(* Logix 5000 project; controller FV vendor 1 type 14 code 217 rev 31.11; software revision 31.00; part 9 of 63 *)
(* tags used below, declared in another part *)
   FR_CFG1_P : PlantItem;   // CFG1_P
   FR_CFG1_P_RawInput : ALIAS FOR RIO_Rack_2:12:I.Data.0;   // FR_CFG1_P
   FR_CFG2_P : PlantItem;   // CFG2_P
   FR_CFG2_P_RawInput : ALIAS FOR RIO_Rack_2:12:I.Data.1;   // FR_CFG2_P
   FR_DEFOAMER : PlantItem;   // DEFOAMER
   FR_DEFOAMER_RawInput : ALIAS FOR RIO_Rack_2:4:I.Data.6;   // FR_DEFOAMER
   FR_Delphi_I : DINT[60];
   FR_FV26_ROTO : PlantItem;   // FV26_ROTO
   FR_FV26_ROTO_RawInput : ALIAS FOR RIO_Rack_2:12:I.Data.10;   // FR_FV26_ROTO
   FR_FV27_ROTO : PlantItem;   // FV27_ROTO
   FR_FV27_ROTO_RawInput : ALIAS FOR RIO_Rack_2:12:I.Data.11;   // FR_FV27_ROTO
   FR_FV28_ROTO : PlantItem;   // FV28_ROTO
   FR_FV28_ROTO_RawInput : ALIAS FOR RIO_Rack_2:12:I.Data.12;   // FR_FV28_ROTO
   FR_FV29_ROTO : PlantItem;   // FV29_ROTO
   FR_FV29_ROTO_RawInput : ALIAS FOR RIO_Rack_2:12:I.Data.13;   // FR_FV29_ROTO
   FR_FV30_ROTO : PlantItem;   // FV30_ROTO
   FR_FV30_ROTO_RawInput : ALIAS FOR RIO_Rack_2:12:I.Data.14;   // FR_FV30_ROTO
   FR_FV31_ROTO : PlantItem;   // FV31_ROTO
   FR_FV31_ROTO_RawInput : ALIAS FOR RIO_Rack_2:12:I.Data.15;   // FR_FV31_ROTO
   FR_OXY_SW1 : PlantItem;   // OXY_SW1
   FR_OXY_SW1_RawInput : ALIAS FOR RIO_Rack_2:3:I.Data.28;   // FR_OXY_SW1
   FR_OXY_SW2 : PlantItem;   // OXY_SW2
   FR_OXY_SW2_RawInput : ALIAS FOR RIO_Rack_2:3:I.Data.29;   // FR_OXY_SW2
   FR_PANELESTOP : PlantItem;   // PANELESTOP
   FR_PANELESTOP_RawInput : ALIAS FOR RIO_Rack_2:3:I.Data.30;   // FR_PANELESTOP
   FR_PARAF : PlantItem;   // PARAF
   FR_PARAF_RawInput : ALIAS FOR RIO_Rack_2:4:I.Data.4;   // FR_PARAF
   FR_PILZ : PlantItem;   // PILZ
   FR_PILZ_RawInput : ALIAS FOR RIO_Rack_2:3:I.Data.31;   // FR_PILZ
   FR_R3_SW3_1 : PlantItem;   // R3_SW3_1
   FR_R3_SW3_1_RawInput : ALIAS FOR RIO_Rack_2:4:I.Data.14;   // FR_R3_SW3_1 FR_N14[109].1
   FR_R3_SW3_2 : PlantItem;   // R3_SW3_2
   FR_R3_SW3_2_RawInput : ALIAS FOR RIO_Rack_2:4:I.Data.10;   // FR_R3_SW3_2 FR_N14[109].0
   FR_YC_IN2 : PlantItem;   // YC_IN2
   FR_YC_IN2_RawInput : ALIAS FOR RIO_Rack_2:12:I.Data.5;   // FR_YC_IN2
   FR_YC_LL : PlantItem;   // YC_LL
   FR_YC_LL_RawInput : ALIAS FOR RIO_Rack_2:12:I.Data.6;   // FR_YC_LL
   One_Second_One_Scan : ALIAS FOR One_Second_1_scan;
(* FR_Common, continued *)

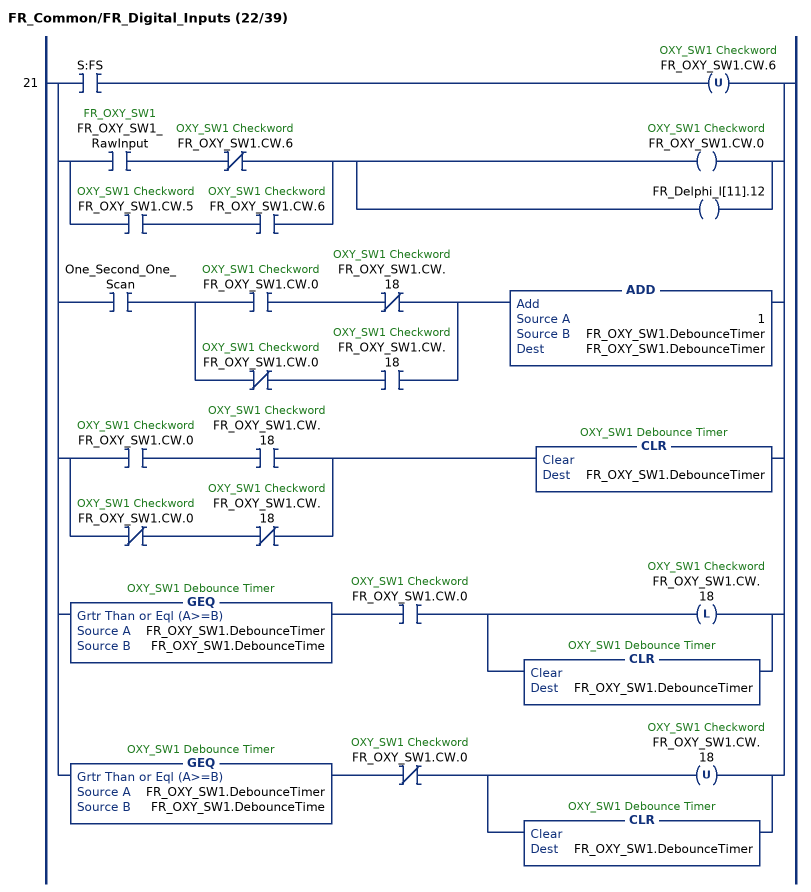
   [picture p94: FR_Common/FR_Digital_Inputs rungs 21-21]
   21: [XIC(S:FS) OTU(FR_OXY_SW1.CW.6) ,[XIC(FR_OXY_SW1_RawInput) XIO(FR_OXY_SW1.CW.6) ,XIC(FR_OXY_SW1.CW.5) XIC(FR_OXY_SW1.CW.6) ] [OTE(FR_OXY_SW1.CW.0) ,OTE(FR_Delphi_I[11].12) ] ,XIC(One_Second_One_Scan) [XIC(FR_OXY_SW1.CW.0) XIO(FR_OXY_SW1.CW.18) ,XIO(FR_OXY_SW1.CW.0) XIC(FR_OXY_SW1.CW.18) ] ADD(1,FR_OXY_SW1.DebounceTimer,FR_OXY_SW1.DebounceTimer) ,[XIC(FR_OXY_SW1.CW.0) XIC(FR_OXY_SW1.CW.18) ,XIO(FR_OXY_SW1.CW.0) XIO(FR_OXY_SW1.CW.18) ] CLR(FR_OXY_SW1.DebounceTimer) ,GEQ(FR_OXY_SW1.DebounceTimer,FR_OXY_SW1.DebounceTime) XIC(FR_OXY_SW1.CW.0) [OTL(FR_OXY_SW1.CW.18) ,CLR(FR_OXY_SW1.DebounceTimer) ] ,GEQ(FR_OXY_SW1.DebounceTimer,FR_OXY_SW1.DebounceTime) XIO(FR_OXY_SW1.CW.0) [OTU(FR_OXY_SW1.CW.18) ,CLR(FR_OXY_SW1.DebounceTimer) ] ];
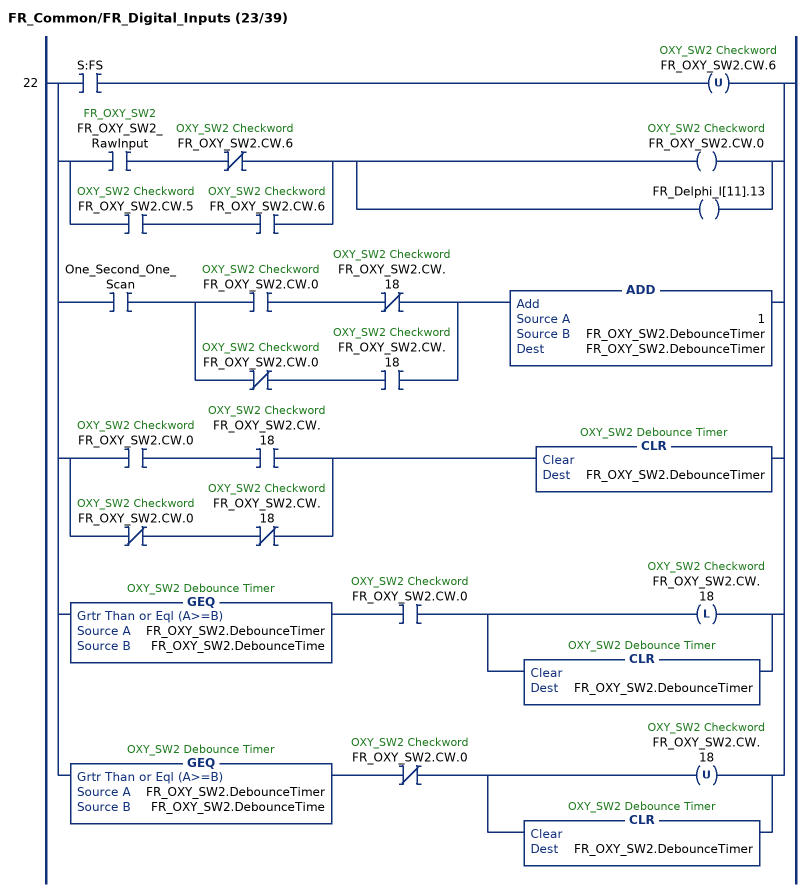
   22: [XIC(S:FS) OTU(FR_OXY_SW2.CW.6) ,[XIC(FR_OXY_SW2_RawInput) XIO(FR_OXY_SW2.CW.6) ,XIC(FR_OXY_SW2.CW.5) XIC(FR_OXY_SW2.CW.6) ] [OTE(FR_OXY_SW2.CW.0) ,OTE(FR_Delphi_I[11].13) ] ,XIC(One_Second_One_Scan) [XIC(FR_OXY_SW2.CW.0) XIO(FR_OXY_SW2.CW.18) ,XIO(FR_OXY_SW2.CW.0) XIC(FR_OXY_SW2.CW.18) ] ADD(1,FR_OXY_SW2.DebounceTimer,FR_OXY_SW2.DebounceTimer) ,[XIC(FR_OXY_SW2.CW.0) XIC(FR_OXY_SW2.CW.18) ,XIO(FR_OXY_SW2.CW.0) XIO(FR_OXY_SW2.CW.18) ] CLR(FR_OXY_SW2.DebounceTimer) ,GEQ(FR_OXY_SW2.DebounceTimer,FR_OXY_SW2.DebounceTime) XIC(FR_OXY_SW2.CW.0) [OTL(FR_OXY_SW2.CW.18) ,CLR(FR_OXY_SW2.DebounceTimer) ] ,GEQ(FR_OXY_SW2.DebounceTimer,FR_OXY_SW2.DebounceTime) XIO(FR_OXY_SW2.CW.0) [OTU(FR_OXY_SW2.CW.18) ,CLR(FR_OXY_SW2.DebounceTimer) ] ];
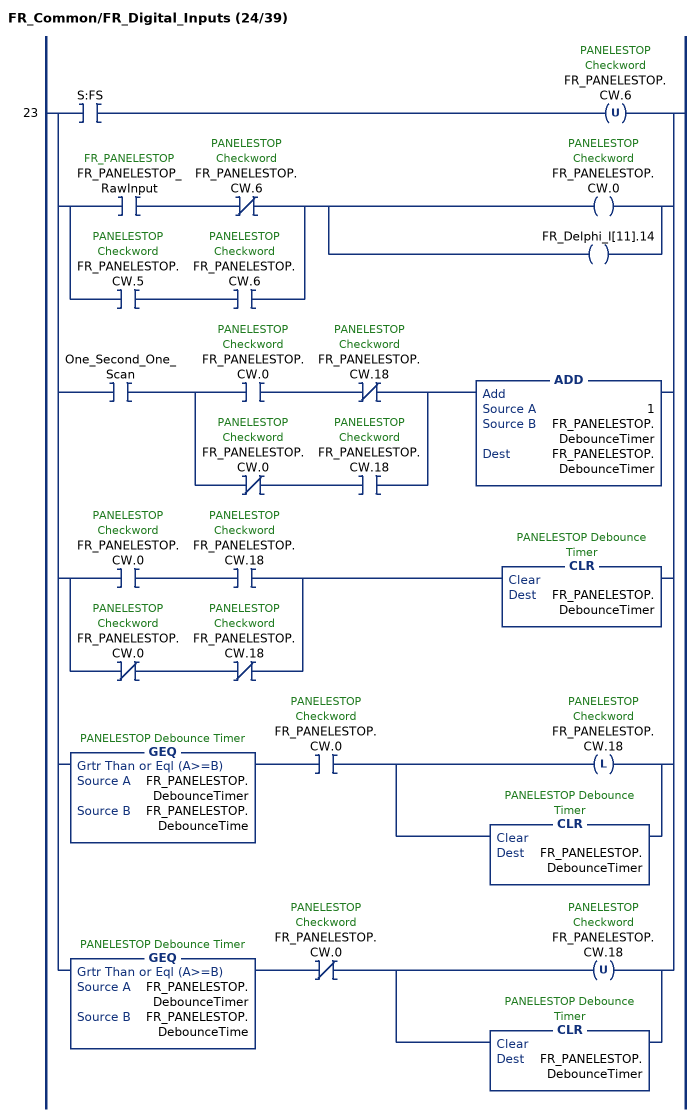
   23: [XIC(S:FS) OTU(FR_PANELESTOP.CW.6) ,[XIC(FR_PANELESTOP_RawInput) XIO(FR_PANELESTOP.CW.6) ,XIC(FR_PANELESTOP.CW.5) XIC(FR_PANELESTOP.CW.6) ] [OTE(FR_PANELESTOP.CW.0) ,OTE(FR_Delphi_I[11].14) ] ,XIC(One_Second_One_Scan) [XIC(FR_PANELESTOP.CW.0) XIO(FR_PANELESTOP.CW.18) ,XIO(FR_PANELESTOP.CW.0) XIC(FR_PANELESTOP.CW.18) ] ADD(1,FR_PANELESTOP.DebounceTimer,FR_PANELESTOP.DebounceTimer) ,[XIC(FR_PANELESTOP.CW.0) XIC(FR_PANELESTOP.CW.18) ,XIO(FR_PANELESTOP.CW.0) XIO(FR_PANELESTOP.CW.18) ] CLR(FR_PANELESTOP.DebounceTimer) ,GEQ(FR_PANELESTOP.DebounceTimer,FR_PANELESTOP.DebounceTime) XIC(FR_PANELESTOP.CW.0) [OTL(FR_PANELESTOP.CW.18) ,CLR(FR_PANELESTOP.DebounceTimer) ] ,GEQ(FR_PANELESTOP.DebounceTimer,FR_PANELESTOP.DebounceTime) XIO(FR_PANELESTOP.CW.0) [OTU(FR_PANELESTOP.CW.18) ,CLR(FR_PANELESTOP.DebounceTimer) ] ];
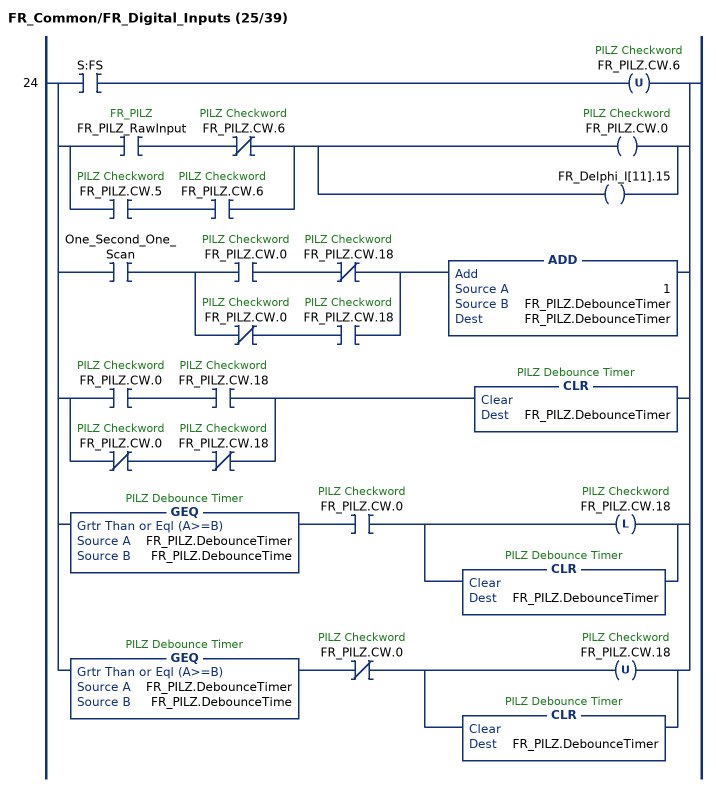
   24: [XIC(S:FS) OTU(FR_PILZ.CW.6) ,[XIC(FR_PILZ_RawInput) XIO(FR_PILZ.CW.6) ,XIC(FR_PILZ.CW.5) XIC(FR_PILZ.CW.6) ] [OTE(FR_PILZ.CW.0) ,OTE(FR_Delphi_I[11].15) ] ,XIC(One_Second_One_Scan) [XIC(FR_PILZ.CW.0) XIO(FR_PILZ.CW.18) ,XIO(FR_PILZ.CW.0) XIC(FR_PILZ.CW.18) ] ADD(1,FR_PILZ.DebounceTimer,FR_PILZ.DebounceTimer) ,[XIC(FR_PILZ.CW.0) XIC(FR_PILZ.CW.18) ,XIO(FR_PILZ.CW.0) XIO(FR_PILZ.CW.18) ] CLR(FR_PILZ.DebounceTimer) ,GEQ(FR_PILZ.DebounceTimer,FR_PILZ.DebounceTime) XIC(FR_PILZ.CW.0) [OTL(FR_PILZ.CW.18) ,CLR(FR_PILZ.DebounceTimer) ] ,GEQ(FR_PILZ.DebounceTimer,FR_PILZ.DebounceTime) XIO(FR_PILZ.CW.0) [OTU(FR_PILZ.CW.18) ,CLR(FR_PILZ.DebounceTimer) ] ];
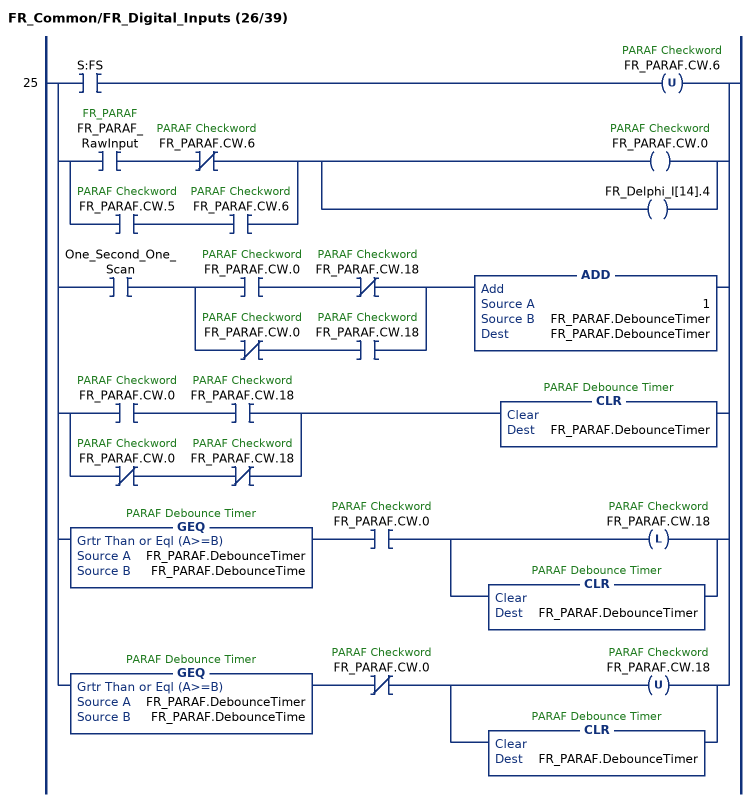
   25: [XIC(S:FS) OTU(FR_PARAF.CW.6) ,[XIC(FR_PARAF_RawInput) XIO(FR_PARAF.CW.6) ,XIC(FR_PARAF.CW.5) XIC(FR_PARAF.CW.6) ] [OTE(FR_PARAF.CW.0) ,OTE(FR_Delphi_I[14].4) ] ,XIC(One_Second_One_Scan) [XIC(FR_PARAF.CW.0) XIO(FR_PARAF.CW.18) ,XIO(FR_PARAF.CW.0) XIC(FR_PARAF.CW.18) ] ADD(1,FR_PARAF.DebounceTimer,FR_PARAF.DebounceTimer) ,[XIC(FR_PARAF.CW.0) XIC(FR_PARAF.CW.18) ,XIO(FR_PARAF.CW.0) XIO(FR_PARAF.CW.18) ] CLR(FR_PARAF.DebounceTimer) ,GEQ(FR_PARAF.DebounceTimer,FR_PARAF.DebounceTime) XIC(FR_PARAF.CW.0) [OTL(FR_PARAF.CW.18) ,CLR(FR_PARAF.DebounceTimer) ] ,GEQ(FR_PARAF.DebounceTimer,FR_PARAF.DebounceTime) XIO(FR_PARAF.CW.0) [OTU(FR_PARAF.CW.18) ,CLR(FR_PARAF.DebounceTimer) ] ];
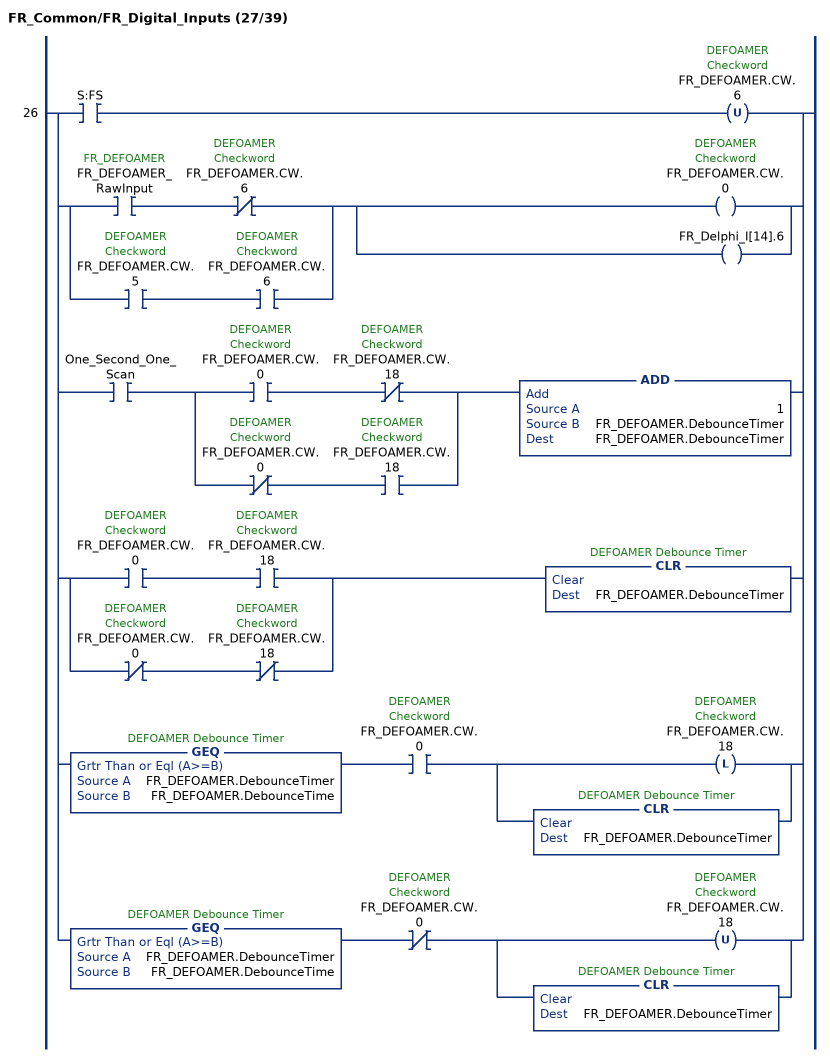
   26: [XIC(S:FS) OTU(FR_DEFOAMER.CW.6) ,[XIC(FR_DEFOAMER_RawInput) XIO(FR_DEFOAMER.CW.6) ,XIC(FR_DEFOAMER.CW.5) XIC(FR_DEFOAMER.CW.6) ] [OTE(FR_DEFOAMER.CW.0) ,OTE(FR_Delphi_I[14].6) ] ,XIC(One_Second_One_Scan) [XIC(FR_DEFOAMER.CW.0) XIO(FR_DEFOAMER.CW.18) ,XIO(FR_DEFOAMER.CW.0) XIC(FR_DEFOAMER.CW.18) ] ADD(1,FR_DEFOAMER.DebounceTimer,FR_DEFOAMER.DebounceTimer) ,[XIC(FR_DEFOAMER.CW.0) XIC(FR_DEFOAMER.CW.18) ,XIO(FR_DEFOAMER.CW.0) XIO(FR_DEFOAMER.CW.18) ] CLR(FR_DEFOAMER.DebounceTimer) ,GEQ(FR_DEFOAMER.DebounceTimer,FR_DEFOAMER.DebounceTime) XIC(FR_DEFOAMER.CW.0) [OTL(FR_DEFOAMER.CW.18) ,CLR(FR_DEFOAMER.DebounceTimer) ] ,GEQ(FR_DEFOAMER.DebounceTimer,FR_DEFOAMER.DebounceTime) XIO(FR_DEFOAMER.CW.0) [OTU(FR_DEFOAMER.CW.18) ,CLR(FR_DEFOAMER.DebounceTimer) ] ];
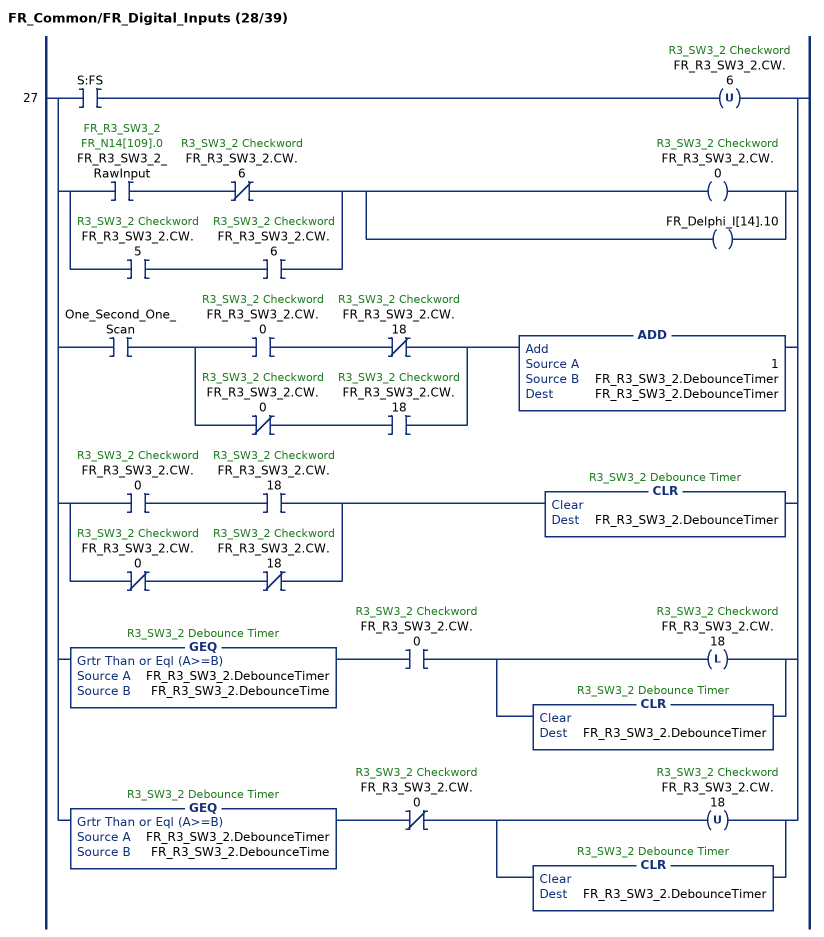
   27: [XIC(S:FS) OTU(FR_R3_SW3_2.CW.6) ,[XIC(FR_R3_SW3_2_RawInput) XIO(FR_R3_SW3_2.CW.6) ,XIC(FR_R3_SW3_2.CW.5) XIC(FR_R3_SW3_2.CW.6) ] [OTE(FR_R3_SW3_2.CW.0) ,OTE(FR_Delphi_I[14].10) ] ,XIC(One_Second_One_Scan) [XIC(FR_R3_SW3_2.CW.0) XIO(FR_R3_SW3_2.CW.18) ,XIO(FR_R3_SW3_2.CW.0) XIC(FR_R3_SW3_2.CW.18) ] ADD(1,FR_R3_SW3_2.DebounceTimer,FR_R3_SW3_2.DebounceTimer) ,[XIC(FR_R3_SW3_2.CW.0) XIC(FR_R3_SW3_2.CW.18) ,XIO(FR_R3_SW3_2.CW.0) XIO(FR_R3_SW3_2.CW.18) ] CLR(FR_R3_SW3_2.DebounceTimer) ,GEQ(FR_R3_SW3_2.DebounceTimer,FR_R3_SW3_2.DebounceTime) XIC(FR_R3_SW3_2.CW.0) [OTL(FR_R3_SW3_2.CW.18) ,CLR(FR_R3_SW3_2.DebounceTimer) ] ,GEQ(FR_R3_SW3_2.DebounceTimer,FR_R3_SW3_2.DebounceTime) XIO(FR_R3_SW3_2.CW.0) [OTU(FR_R3_SW3_2.CW.18) ,CLR(FR_R3_SW3_2.DebounceTimer) ] ];
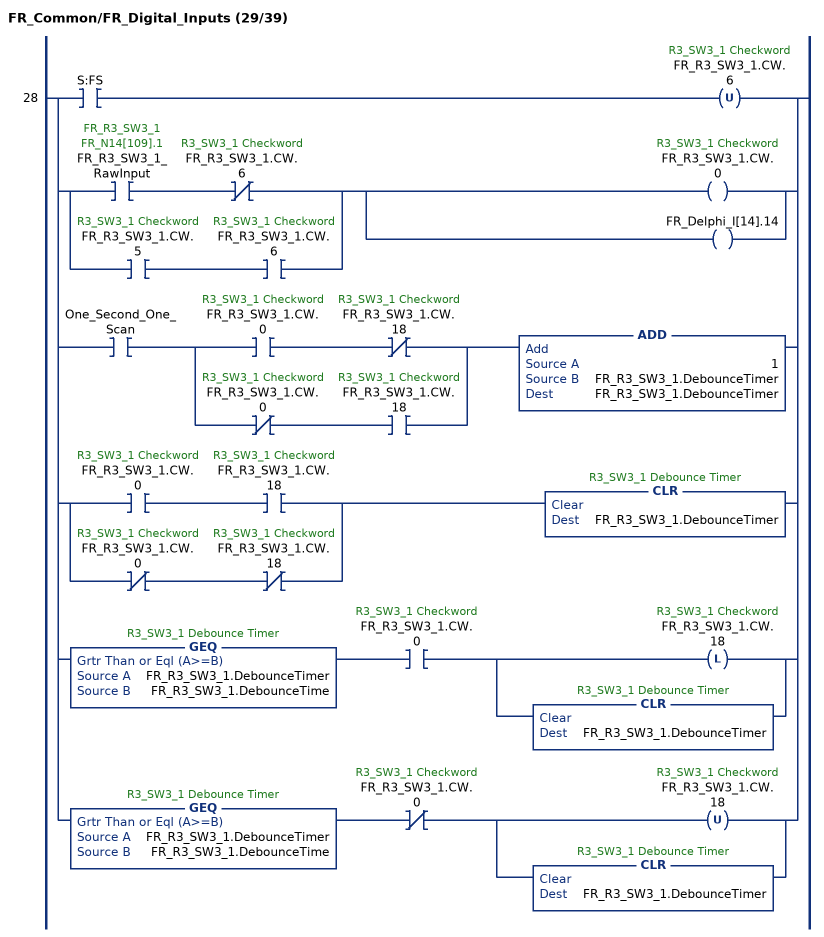
   28: [XIC(S:FS) OTU(FR_R3_SW3_1.CW.6) ,[XIC(FR_R3_SW3_1_RawInput) XIO(FR_R3_SW3_1.CW.6) ,XIC(FR_R3_SW3_1.CW.5) XIC(FR_R3_SW3_1.CW.6) ] [OTE(FR_R3_SW3_1.CW.0) ,OTE(FR_Delphi_I[14].14) ] ,XIC(One_Second_One_Scan) [XIC(FR_R3_SW3_1.CW.0) XIO(FR_R3_SW3_1.CW.18) ,XIO(FR_R3_SW3_1.CW.0) XIC(FR_R3_SW3_1.CW.18) ] ADD(1,FR_R3_SW3_1.DebounceTimer,FR_R3_SW3_1.DebounceTimer) ,[XIC(FR_R3_SW3_1.CW.0) XIC(FR_R3_SW3_1.CW.18) ,XIO(FR_R3_SW3_1.CW.0) XIO(FR_R3_SW3_1.CW.18) ] CLR(FR_R3_SW3_1.DebounceTimer) ,GEQ(FR_R3_SW3_1.DebounceTimer,FR_R3_SW3_1.DebounceTime) XIC(FR_R3_SW3_1.CW.0) [OTL(FR_R3_SW3_1.CW.18) ,CLR(FR_R3_SW3_1.DebounceTimer) ] ,GEQ(FR_R3_SW3_1.DebounceTimer,FR_R3_SW3_1.DebounceTime) XIO(FR_R3_SW3_1.CW.0) [OTU(FR_R3_SW3_1.CW.18) ,CLR(FR_R3_SW3_1.DebounceTimer) ] ];
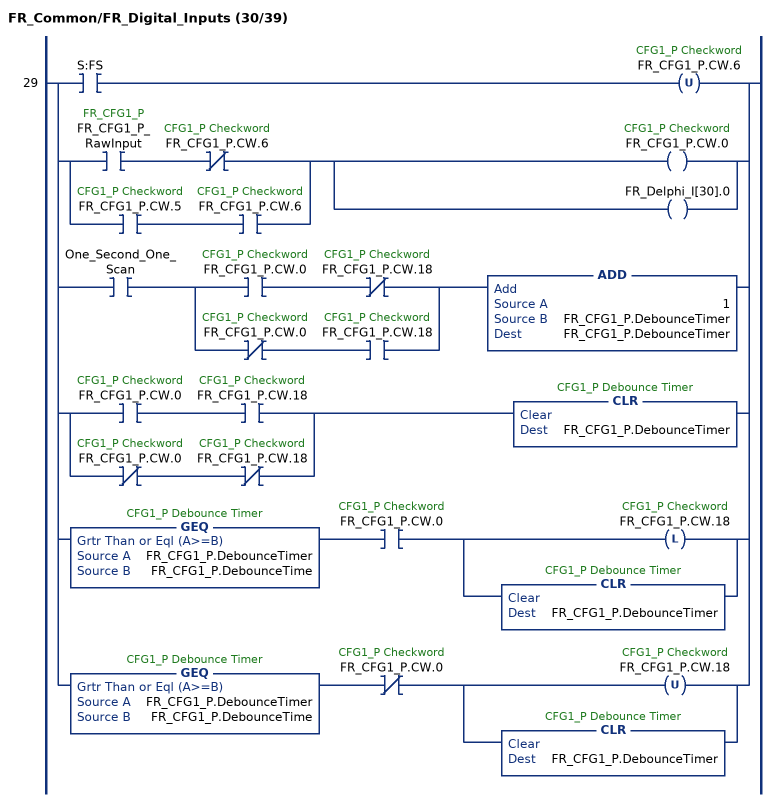
   29: [XIC(S:FS) OTU(FR_CFG1_P.CW.6) ,[XIC(FR_CFG1_P_RawInput) XIO(FR_CFG1_P.CW.6) ,XIC(FR_CFG1_P.CW.5) XIC(FR_CFG1_P.CW.6) ] [OTE(FR_CFG1_P.CW.0) ,OTE(FR_Delphi_I[30].0) ] ,XIC(One_Second_One_Scan) [XIC(FR_CFG1_P.CW.0) XIO(FR_CFG1_P.CW.18) ,XIO(FR_CFG1_P.CW.0) XIC(FR_CFG1_P.CW.18) ] ADD(1,FR_CFG1_P.DebounceTimer,FR_CFG1_P.DebounceTimer) ,[XIC(FR_CFG1_P.CW.0) XIC(FR_CFG1_P.CW.18) ,XIO(FR_CFG1_P.CW.0) XIO(FR_CFG1_P.CW.18) ] CLR(FR_CFG1_P.DebounceTimer) ,GEQ(FR_CFG1_P.DebounceTimer,FR_CFG1_P.DebounceTime) XIC(FR_CFG1_P.CW.0) [OTL(FR_CFG1_P.CW.18) ,CLR(FR_CFG1_P.DebounceTimer) ] ,GEQ(FR_CFG1_P.DebounceTimer,FR_CFG1_P.DebounceTime) XIO(FR_CFG1_P.CW.0) [OTU(FR_CFG1_P.CW.18) ,CLR(FR_CFG1_P.DebounceTimer) ] ];
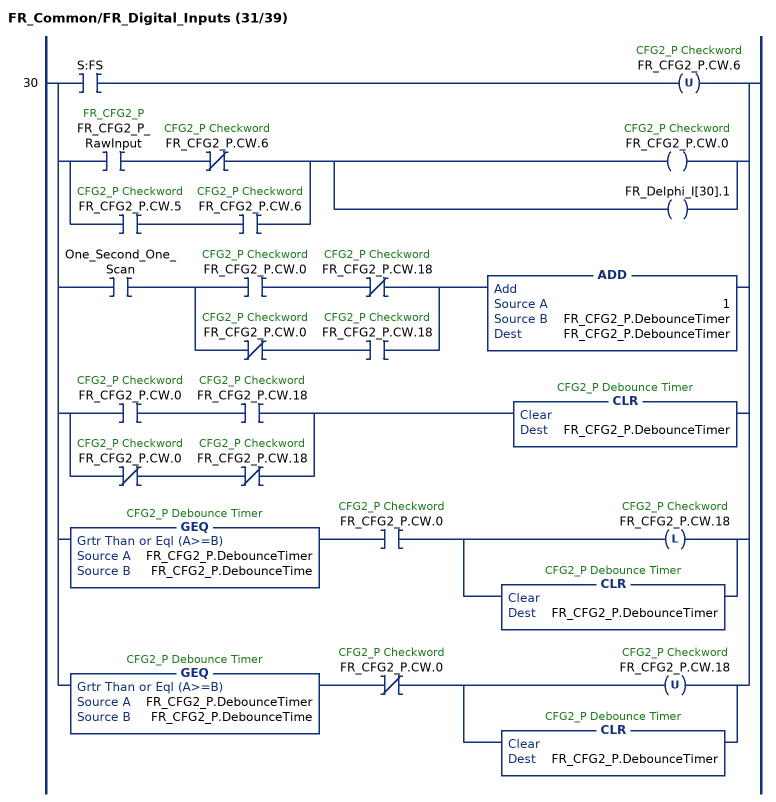
   30: [XIC(S:FS) OTU(FR_CFG2_P.CW.6) ,[XIC(FR_CFG2_P_RawInput) XIO(FR_CFG2_P.CW.6) ,XIC(FR_CFG2_P.CW.5) XIC(FR_CFG2_P.CW.6) ] [OTE(FR_CFG2_P.CW.0) ,OTE(FR_Delphi_I[30].1) ] ,XIC(One_Second_One_Scan) [XIC(FR_CFG2_P.CW.0) XIO(FR_CFG2_P.CW.18) ,XIO(FR_CFG2_P.CW.0) XIC(FR_CFG2_P.CW.18) ] ADD(1,FR_CFG2_P.DebounceTimer,FR_CFG2_P.DebounceTimer) ,[XIC(FR_CFG2_P.CW.0) XIC(FR_CFG2_P.CW.18) ,XIO(FR_CFG2_P.CW.0) XIO(FR_CFG2_P.CW.18) ] CLR(FR_CFG2_P.DebounceTimer) ,GEQ(FR_CFG2_P.DebounceTimer,FR_CFG2_P.DebounceTime) XIC(FR_CFG2_P.CW.0) [OTL(FR_CFG2_P.CW.18) ,CLR(FR_CFG2_P.DebounceTimer) ] ,GEQ(FR_CFG2_P.DebounceTimer,FR_CFG2_P.DebounceTime) XIO(FR_CFG2_P.CW.0) [OTU(FR_CFG2_P.CW.18) ,CLR(FR_CFG2_P.DebounceTimer) ] ];
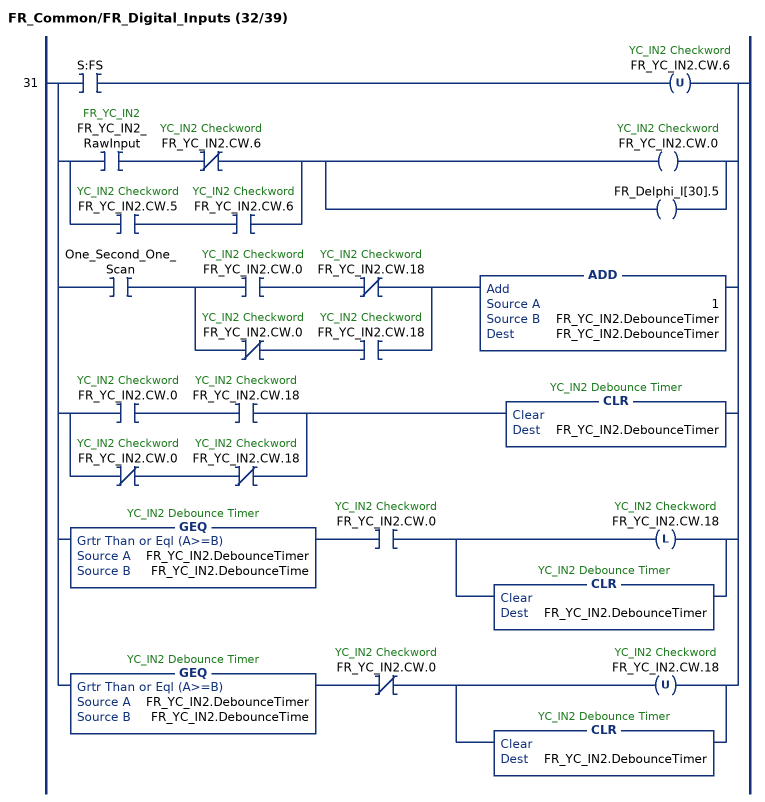
   31: [XIC(S:FS) OTU(FR_YC_IN2.CW.6) ,[XIC(FR_YC_IN2_RawInput) XIO(FR_YC_IN2.CW.6) ,XIC(FR_YC_IN2.CW.5) XIC(FR_YC_IN2.CW.6) ] [OTE(FR_YC_IN2.CW.0) ,OTE(FR_Delphi_I[30].5) ] ,XIC(One_Second_One_Scan) [XIC(FR_YC_IN2.CW.0) XIO(FR_YC_IN2.CW.18) ,XIO(FR_YC_IN2.CW.0) XIC(FR_YC_IN2.CW.18) ] ADD(1,FR_YC_IN2.DebounceTimer,FR_YC_IN2.DebounceTimer) ,[XIC(FR_YC_IN2.CW.0) XIC(FR_YC_IN2.CW.18) ,XIO(FR_YC_IN2.CW.0) XIO(FR_YC_IN2.CW.18) ] CLR(FR_YC_IN2.DebounceTimer) ,GEQ(FR_YC_IN2.DebounceTimer,FR_YC_IN2.DebounceTime) XIC(FR_YC_IN2.CW.0) [OTL(FR_YC_IN2.CW.18) ,CLR(FR_YC_IN2.DebounceTimer) ] ,GEQ(FR_YC_IN2.DebounceTimer,FR_YC_IN2.DebounceTime) XIO(FR_YC_IN2.CW.0) [OTU(FR_YC_IN2.CW.18) ,CLR(FR_YC_IN2.DebounceTimer) ] ];
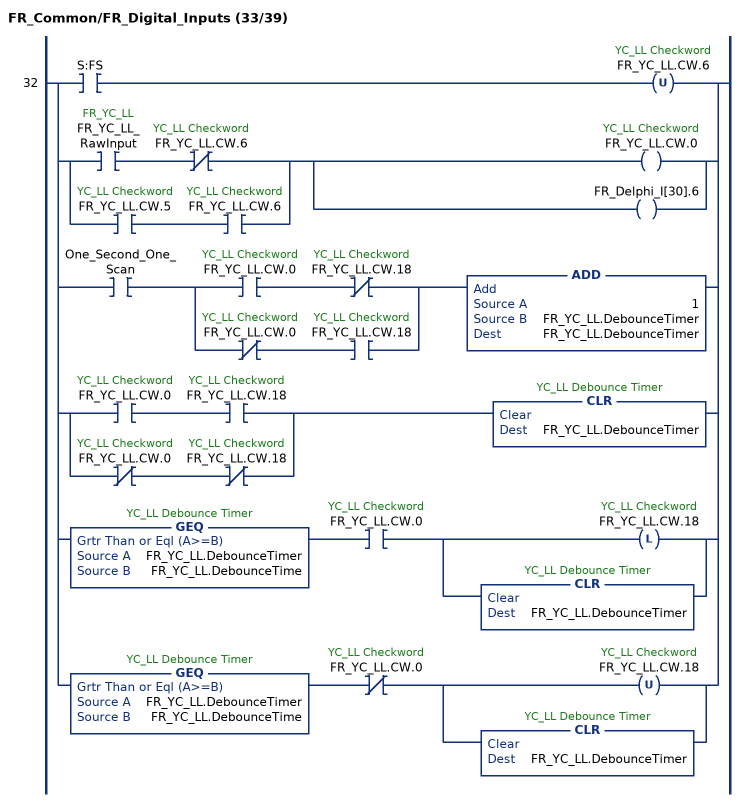
   32: [XIC(S:FS) OTU(FR_YC_LL.CW.6) ,[XIC(FR_YC_LL_RawInput) XIO(FR_YC_LL.CW.6) ,XIC(FR_YC_LL.CW.5) XIC(FR_YC_LL.CW.6) ] [OTE(FR_YC_LL.CW.0) ,OTE(FR_Delphi_I[30].6) ] ,XIC(One_Second_One_Scan) [XIC(FR_YC_LL.CW.0) XIO(FR_YC_LL.CW.18) ,XIO(FR_YC_LL.CW.0) XIC(FR_YC_LL.CW.18) ] ADD(1,FR_YC_LL.DebounceTimer,FR_YC_LL.DebounceTimer) ,[XIC(FR_YC_LL.CW.0) XIC(FR_YC_LL.CW.18) ,XIO(FR_YC_LL.CW.0) XIO(FR_YC_LL.CW.18) ] CLR(FR_YC_LL.DebounceTimer) ,GEQ(FR_YC_LL.DebounceTimer,FR_YC_LL.DebounceTime) XIC(FR_YC_LL.CW.0) [OTL(FR_YC_LL.CW.18) ,CLR(FR_YC_LL.DebounceTimer) ] ,GEQ(FR_YC_LL.DebounceTimer,FR_YC_LL.DebounceTime) XIO(FR_YC_LL.CW.0) [OTU(FR_YC_LL.CW.18) ,CLR(FR_YC_LL.DebounceTimer) ] ];
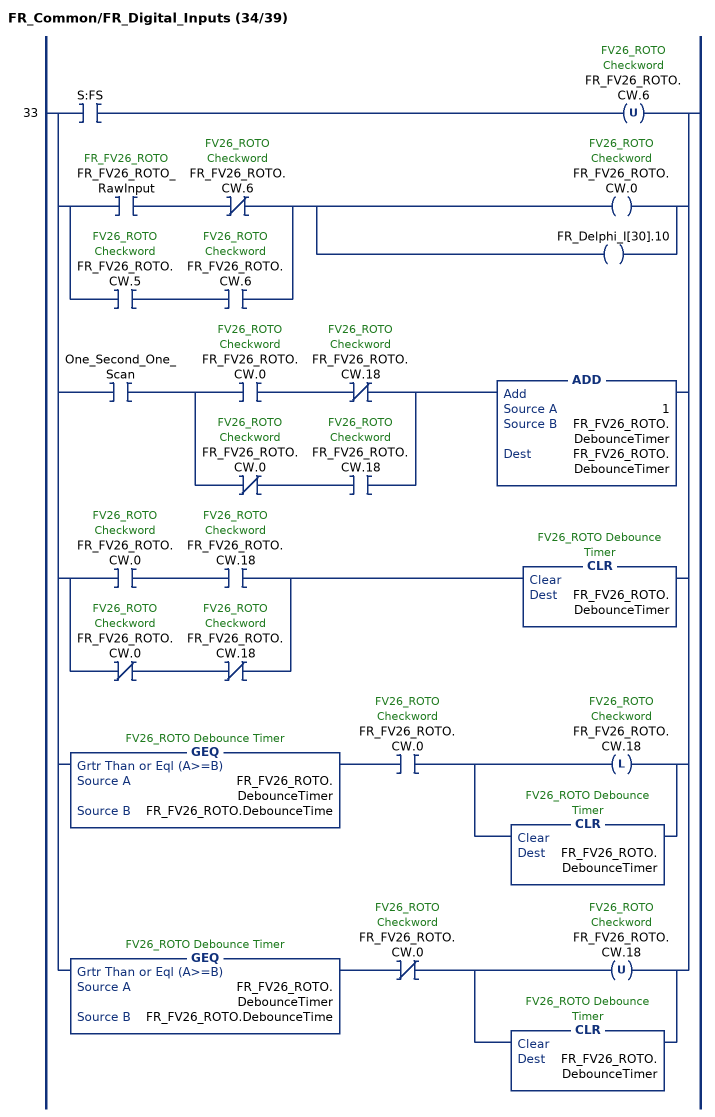
   33: [XIC(S:FS) OTU(FR_FV26_ROTO.CW.6) ,[XIC(FR_FV26_ROTO_RawInput) XIO(FR_FV26_ROTO.CW.6) ,XIC(FR_FV26_ROTO.CW.5) XIC(FR_FV26_ROTO.CW.6) ] [OTE(FR_FV26_ROTO.CW.0) ,OTE(FR_Delphi_I[30].10) ] ,XIC(One_Second_One_Scan) [XIC(FR_FV26_ROTO.CW.0) XIO(FR_FV26_ROTO.CW.18) ,XIO(FR_FV26_ROTO.CW.0) XIC(FR_FV26_ROTO.CW.18) ] ADD(1,FR_FV26_ROTO.DebounceTimer,FR_FV26_ROTO.DebounceTimer) ,[XIC(FR_FV26_ROTO.CW.0) XIC(FR_FV26_ROTO.CW.18) ,XIO(FR_FV26_ROTO.CW.0) XIO(FR_FV26_ROTO.CW.18) ] CLR(FR_FV26_ROTO.DebounceTimer) ,GEQ(FR_FV26_ROTO.DebounceTimer,FR_FV26_ROTO.DebounceTime) XIC(FR_FV26_ROTO.CW.0) [OTL(FR_FV26_ROTO.CW.18) ,CLR(FR_FV26_ROTO.DebounceTimer) ] ,GEQ(FR_FV26_ROTO.DebounceTimer,FR_FV26_ROTO.DebounceTime) XIO(FR_FV26_ROTO.CW.0) [OTU(FR_FV26_ROTO.CW.18) ,CLR(FR_FV26_ROTO.DebounceTimer) ] ];
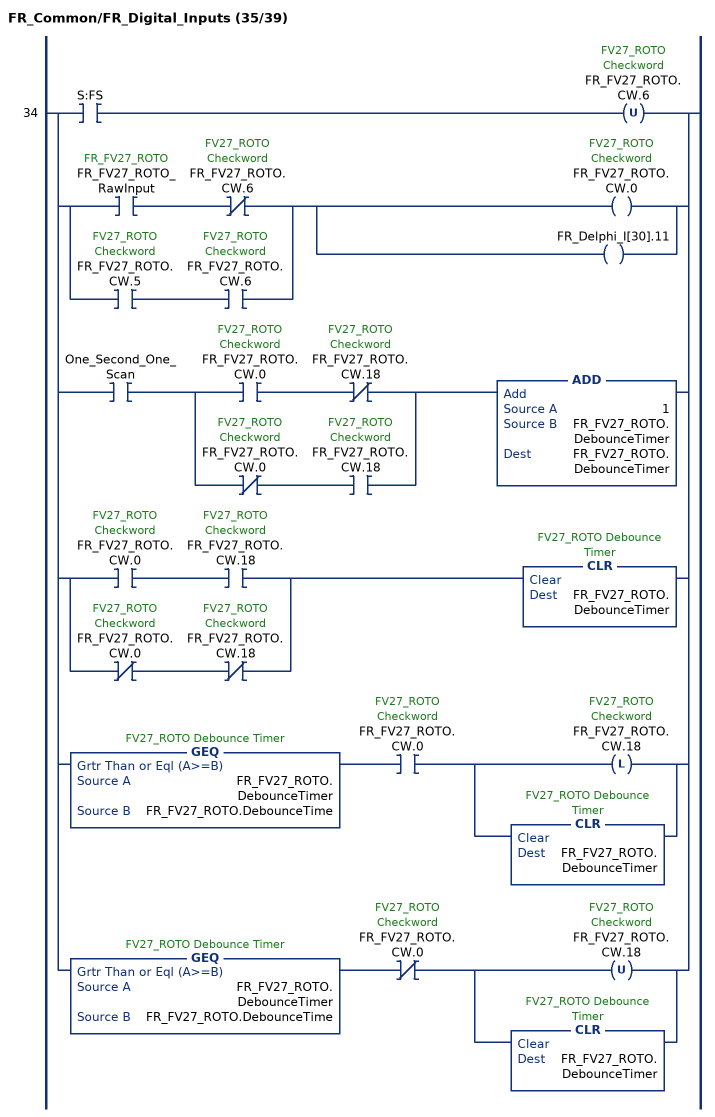
   34: [XIC(S:FS) OTU(FR_FV27_ROTO.CW.6) ,[XIC(FR_FV27_ROTO_RawInput) XIO(FR_FV27_ROTO.CW.6) ,XIC(FR_FV27_ROTO.CW.5) XIC(FR_FV27_ROTO.CW.6) ] [OTE(FR_FV27_ROTO.CW.0) ,OTE(FR_Delphi_I[30].11) ] ,XIC(One_Second_One_Scan) [XIC(FR_FV27_ROTO.CW.0) XIO(FR_FV27_ROTO.CW.18) ,XIO(FR_FV27_ROTO.CW.0) XIC(FR_FV27_ROTO.CW.18) ] ADD(1,FR_FV27_ROTO.DebounceTimer,FR_FV27_ROTO.DebounceTimer) ,[XIC(FR_FV27_ROTO.CW.0) XIC(FR_FV27_ROTO.CW.18) ,XIO(FR_FV27_ROTO.CW.0) XIO(FR_FV27_ROTO.CW.18) ] CLR(FR_FV27_ROTO.DebounceTimer) ,GEQ(FR_FV27_ROTO.DebounceTimer,FR_FV27_ROTO.DebounceTime) XIC(FR_FV27_ROTO.CW.0) [OTL(FR_FV27_ROTO.CW.18) ,CLR(FR_FV27_ROTO.DebounceTimer) ] ,GEQ(FR_FV27_ROTO.DebounceTimer,FR_FV27_ROTO.DebounceTime) XIO(FR_FV27_ROTO.CW.0) [OTU(FR_FV27_ROTO.CW.18) ,CLR(FR_FV27_ROTO.DebounceTimer) ] ];
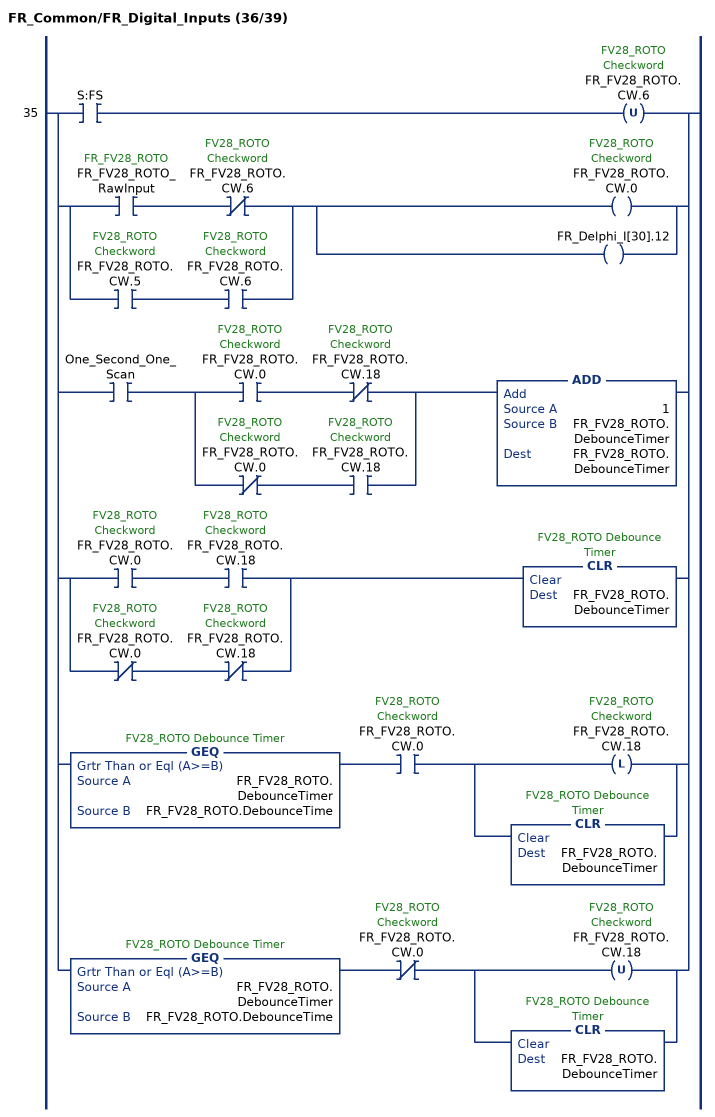
   35: [XIC(S:FS) OTU(FR_FV28_ROTO.CW.6) ,[XIC(FR_FV28_ROTO_RawInput) XIO(FR_FV28_ROTO.CW.6) ,XIC(FR_FV28_ROTO.CW.5) XIC(FR_FV28_ROTO.CW.6) ] [OTE(FR_FV28_ROTO.CW.0) ,OTE(FR_Delphi_I[30].12) ] ,XIC(One_Second_One_Scan) [XIC(FR_FV28_ROTO.CW.0) XIO(FR_FV28_ROTO.CW.18) ,XIO(FR_FV28_ROTO.CW.0) XIC(FR_FV28_ROTO.CW.18) ] ADD(1,FR_FV28_ROTO.DebounceTimer,FR_FV28_ROTO.DebounceTimer) ,[XIC(FR_FV28_ROTO.CW.0) XIC(FR_FV28_ROTO.CW.18) ,XIO(FR_FV28_ROTO.CW.0) XIO(FR_FV28_ROTO.CW.18) ] CLR(FR_FV28_ROTO.DebounceTimer) ,GEQ(FR_FV28_ROTO.DebounceTimer,FR_FV28_ROTO.DebounceTime) XIC(FR_FV28_ROTO.CW.0) [OTL(FR_FV28_ROTO.CW.18) ,CLR(FR_FV28_ROTO.DebounceTimer) ] ,GEQ(FR_FV28_ROTO.DebounceTimer,FR_FV28_ROTO.DebounceTime) XIO(FR_FV28_ROTO.CW.0) [OTU(FR_FV28_ROTO.CW.18) ,CLR(FR_FV28_ROTO.DebounceTimer) ] ];
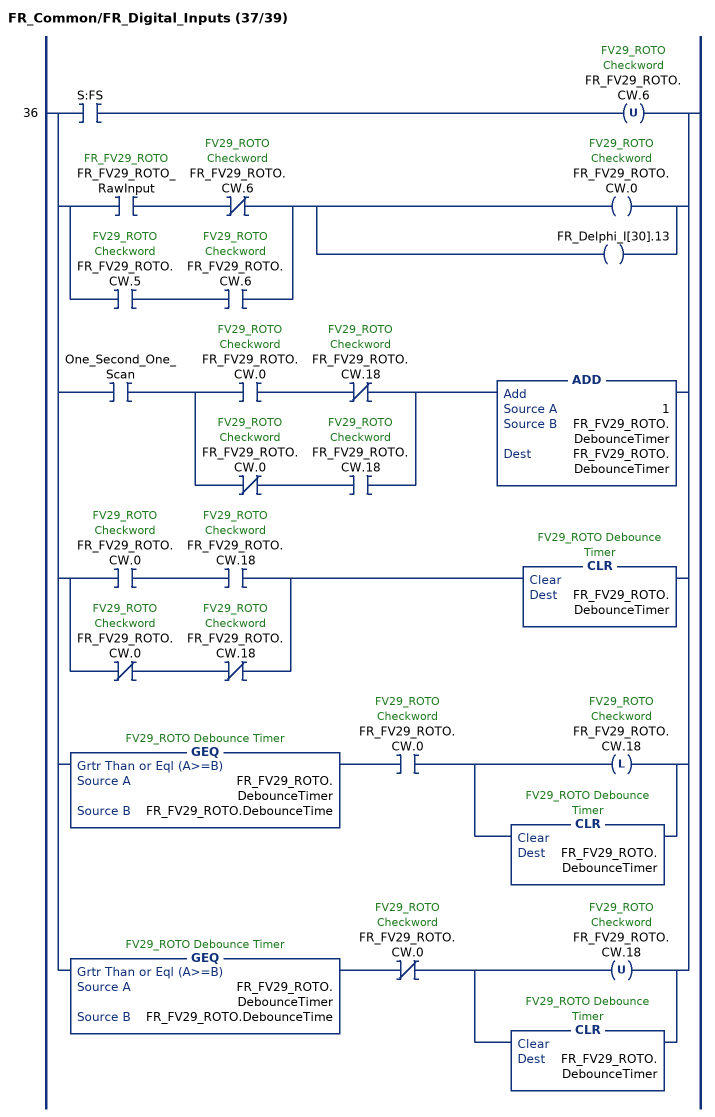
   36: [XIC(S:FS) OTU(FR_FV29_ROTO.CW.6) ,[XIC(FR_FV29_ROTO_RawInput) XIO(FR_FV29_ROTO.CW.6) ,XIC(FR_FV29_ROTO.CW.5) XIC(FR_FV29_ROTO.CW.6) ] [OTE(FR_FV29_ROTO.CW.0) ,OTE(FR_Delphi_I[30].13) ] ,XIC(One_Second_One_Scan) [XIC(FR_FV29_ROTO.CW.0) XIO(FR_FV29_ROTO.CW.18) ,XIO(FR_FV29_ROTO.CW.0) XIC(FR_FV29_ROTO.CW.18) ] ADD(1,FR_FV29_ROTO.DebounceTimer,FR_FV29_ROTO.DebounceTimer) ,[XIC(FR_FV29_ROTO.CW.0) XIC(FR_FV29_ROTO.CW.18) ,XIO(FR_FV29_ROTO.CW.0) XIO(FR_FV29_ROTO.CW.18) ] CLR(FR_FV29_ROTO.DebounceTimer) ,GEQ(FR_FV29_ROTO.DebounceTimer,FR_FV29_ROTO.DebounceTime) XIC(FR_FV29_ROTO.CW.0) [OTL(FR_FV29_ROTO.CW.18) ,CLR(FR_FV29_ROTO.DebounceTimer) ] ,GEQ(FR_FV29_ROTO.DebounceTimer,FR_FV29_ROTO.DebounceTime) XIO(FR_FV29_ROTO.CW.0) [OTU(FR_FV29_ROTO.CW.18) ,CLR(FR_FV29_ROTO.DebounceTimer) ] ];
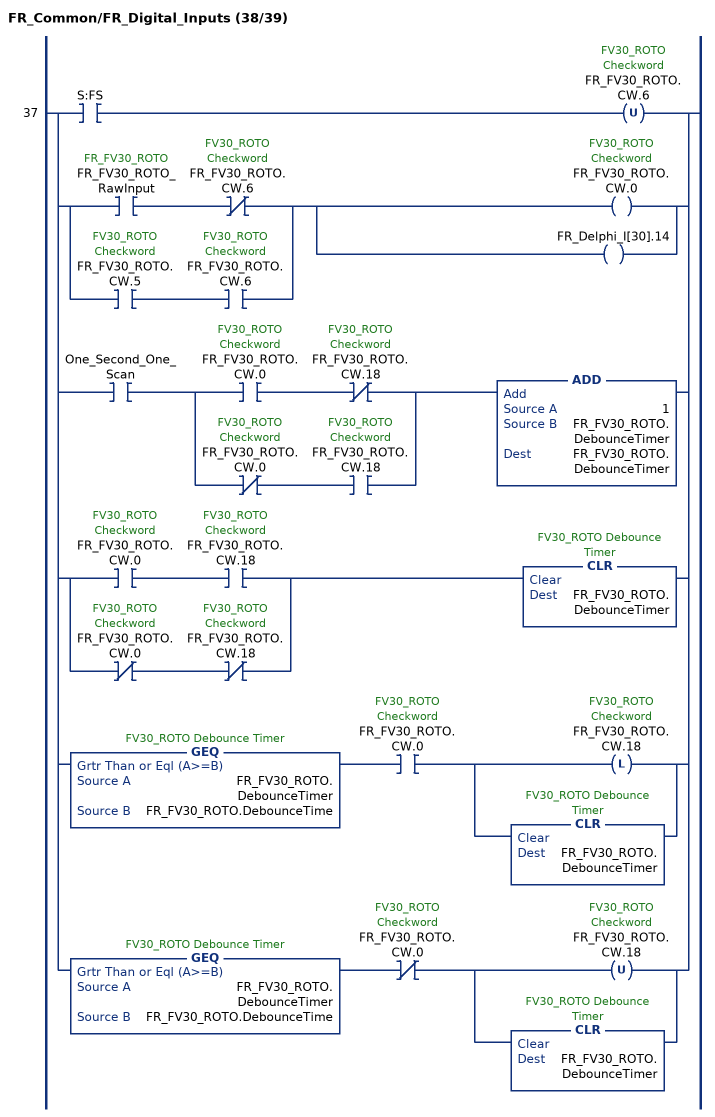
   37: [XIC(S:FS) OTU(FR_FV30_ROTO.CW.6) ,[XIC(FR_FV30_ROTO_RawInput) XIO(FR_FV30_ROTO.CW.6) ,XIC(FR_FV30_ROTO.CW.5) XIC(FR_FV30_ROTO.CW.6) ] [OTE(FR_FV30_ROTO.CW.0) ,OTE(FR_Delphi_I[30].14) ] ,XIC(One_Second_One_Scan) [XIC(FR_FV30_ROTO.CW.0) XIO(FR_FV30_ROTO.CW.18) ,XIO(FR_FV30_ROTO.CW.0) XIC(FR_FV30_ROTO.CW.18) ] ADD(1,FR_FV30_ROTO.DebounceTimer,FR_FV30_ROTO.DebounceTimer) ,[XIC(FR_FV30_ROTO.CW.0) XIC(FR_FV30_ROTO.CW.18) ,XIO(FR_FV30_ROTO.CW.0) XIO(FR_FV30_ROTO.CW.18) ] CLR(FR_FV30_ROTO.DebounceTimer) ,GEQ(FR_FV30_ROTO.DebounceTimer,FR_FV30_ROTO.DebounceTime) XIC(FR_FV30_ROTO.CW.0) [OTL(FR_FV30_ROTO.CW.18) ,CLR(FR_FV30_ROTO.DebounceTimer) ] ,GEQ(FR_FV30_ROTO.DebounceTimer,FR_FV30_ROTO.DebounceTime) XIO(FR_FV30_ROTO.CW.0) [OTU(FR_FV30_ROTO.CW.18) ,CLR(FR_FV30_ROTO.DebounceTimer) ] ];
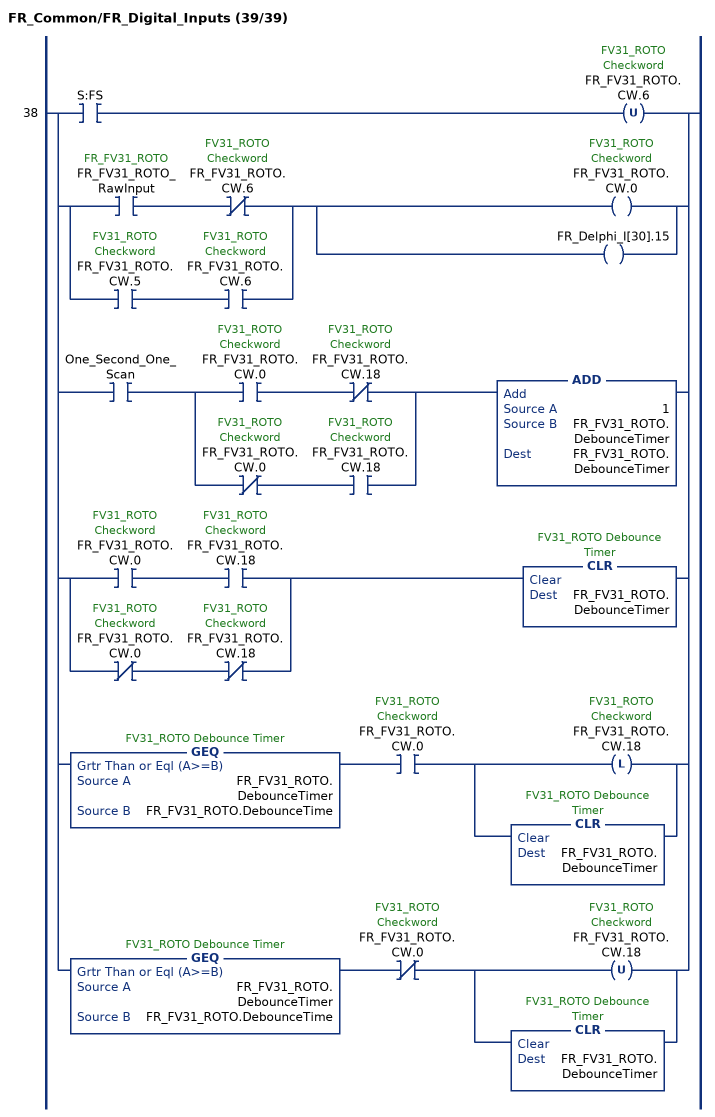
   38: [XIC(S:FS) OTU(FR_FV31_ROTO.CW.6) ,[XIC(FR_FV31_ROTO_RawInput) XIO(FR_FV31_ROTO.CW.6) ,XIC(FR_FV31_ROTO.CW.5) XIC(FR_FV31_ROTO.CW.6) ] [OTE(FR_FV31_ROTO.CW.0) ,OTE(FR_Delphi_I[30].15) ] ,XIC(One_Second_One_Scan) [XIC(FR_FV31_ROTO.CW.0) XIO(FR_FV31_ROTO.CW.18) ,XIO(FR_FV31_ROTO.CW.0) XIC(FR_FV31_ROTO.CW.18) ] ADD(1,FR_FV31_ROTO.DebounceTimer,FR_FV31_ROTO.DebounceTimer) ,[XIC(FR_FV31_ROTO.CW.0) XIC(FR_FV31_ROTO.CW.18) ,XIO(FR_FV31_ROTO.CW.0) XIO(FR_FV31_ROTO.CW.18) ] CLR(FR_FV31_ROTO.DebounceTimer) ,GEQ(FR_FV31_ROTO.DebounceTimer,FR_FV31_ROTO.DebounceTime) XIC(FR_FV31_ROTO.CW.0) [OTL(FR_FV31_ROTO.CW.18) ,CLR(FR_FV31_ROTO.DebounceTimer) ] ,GEQ(FR_FV31_ROTO.DebounceTimer,FR_FV31_ROTO.DebounceTime) XIO(FR_FV31_ROTO.CW.0) [OTU(FR_FV31_ROTO.CW.18) ,CLR(FR_FV31_ROTO.DebounceTimer) ] ];
END_ROUTINE
